// TIA Portal project "TestEssProtoFreia" (V13) (continued)
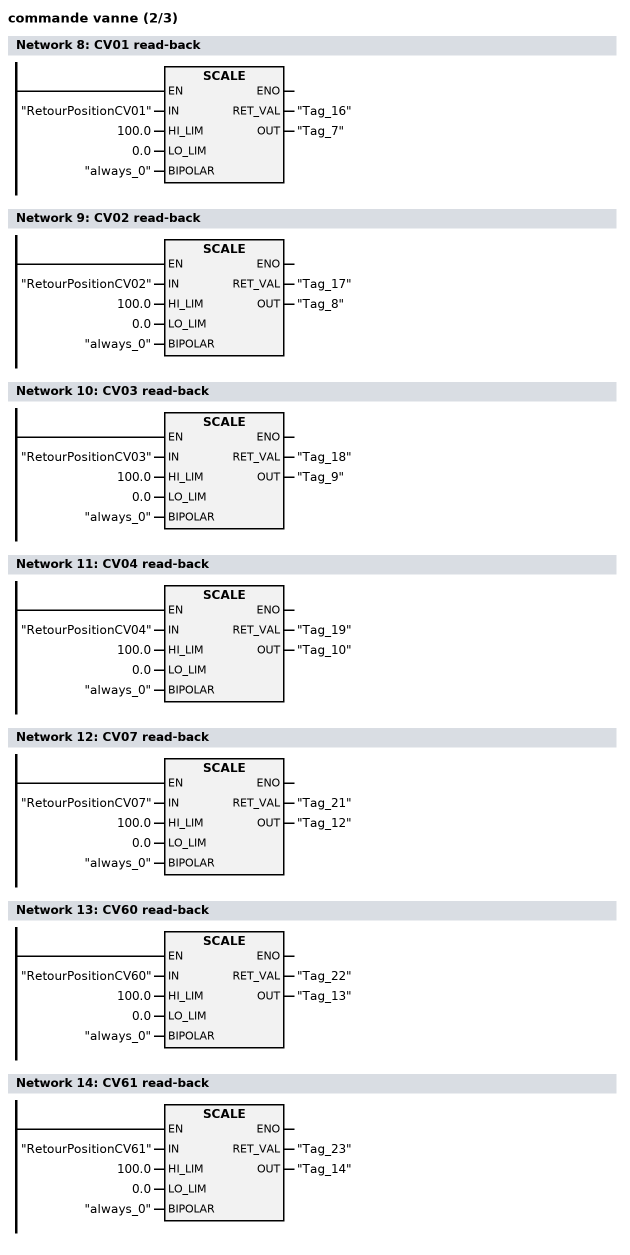
   "Tag_16" := SCALE(IN := "RetourPositionCV01",
                     HI_LIM := 100.0,
                     LO_LIM := 0.0,
                     BIPOLAR := "always_0",
                     OUT => "Tag_7");
END_REGION

REGION Network 9: CV02 read-back
   "Tag_17" := SCALE(IN := "RetourPositionCV02",
                     HI_LIM := 100.0,
                     LO_LIM := 0.0,
                     BIPOLAR := "always_0",
                     OUT => "Tag_8");
END_REGION

REGION Network 10: CV03 read-back
   "Tag_18" := SCALE(IN := "RetourPositionCV03",
                     HI_LIM := 100.0,
                     LO_LIM := 0.0,
                     BIPOLAR := "always_0",
                     OUT => "Tag_9");
END_REGION

REGION Network 11: CV04 read-back
   "Tag_19" := SCALE(IN := "RetourPositionCV04",
                     HI_LIM := 100.0,
                     LO_LIM := 0.0,
                     BIPOLAR := "always_0",
                     OUT => "Tag_10");
END_REGION

REGION Network 12: CV07 read-back
   "Tag_21" := SCALE(IN := "RetourPositionCV07",
                     HI_LIM := 100.0,
                     LO_LIM := 0.0,
                     BIPOLAR := "always_0",
                     OUT => "Tag_12");
END_REGION

REGION Network 13: CV60 read-back
   "Tag_22" := SCALE(IN := "RetourPositionCV60",
                     HI_LIM := 100.0,
                     LO_LIM := 0.0,
                     BIPOLAR := "always_0",
                     OUT => "Tag_13");
END_REGION

REGION Network 14: CV61 read-back
   "Tag_23" := SCALE(IN := "RetourPositionCV61",
                     HI_LIM := 100.0,
                     LO_LIM := 0.0,
                     BIPOLAR := "always_0",
                     OUT => "Tag_14");
END_REGION

REGION Network 15: activation PID CV03 LT03>=80%
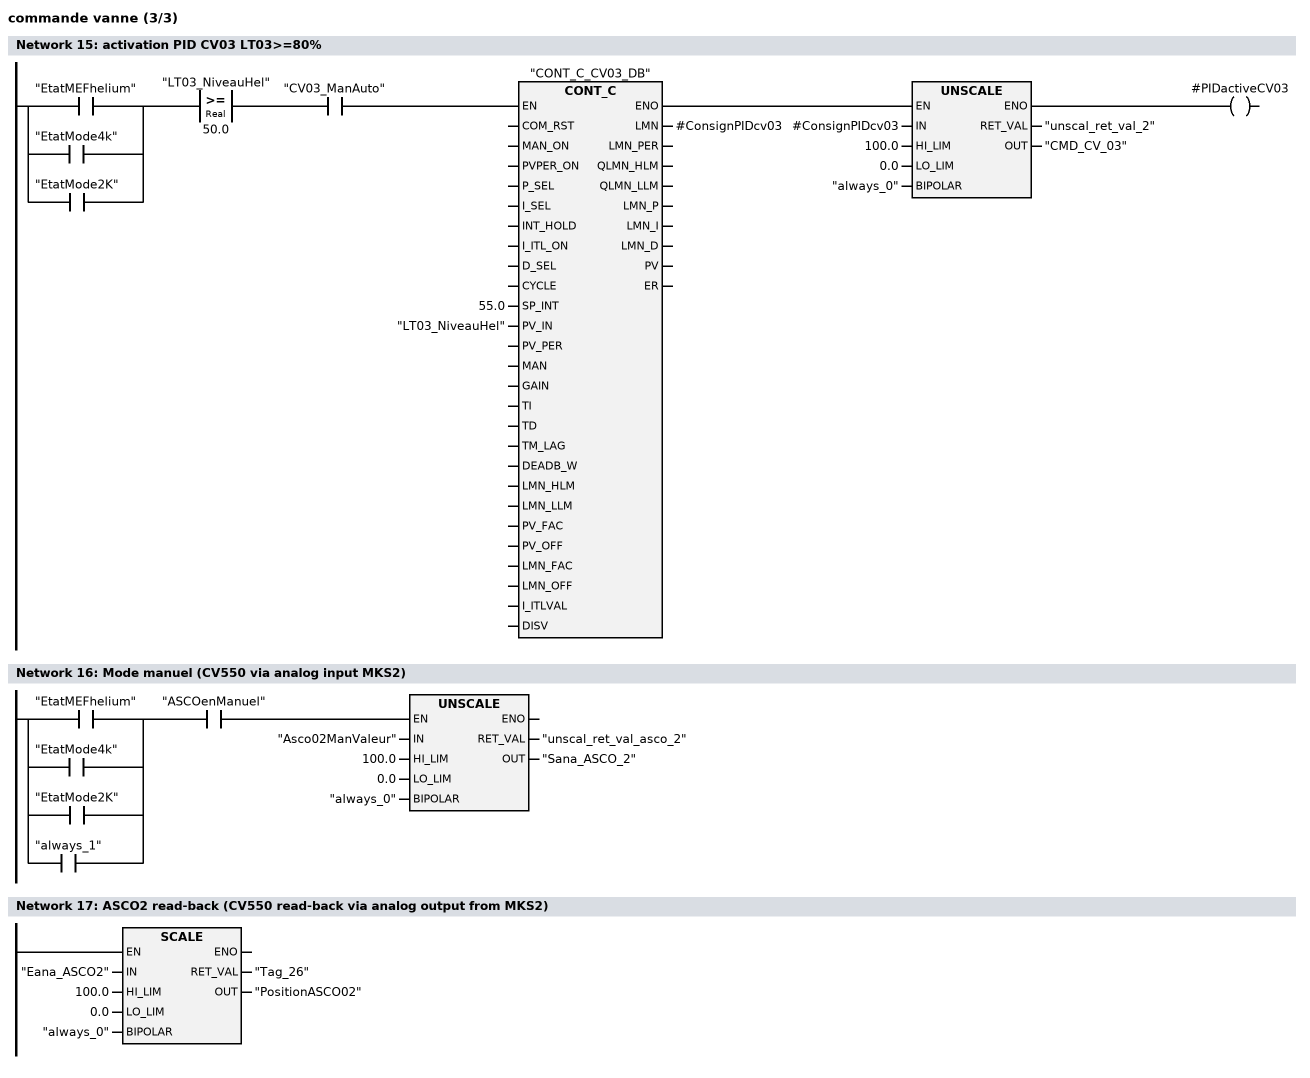
   // ENO of a box is taken as its EN; it also drops when the box reports an error
   #_w1 := ("EtatMEFhelium" OR "EtatMode4k" OR "EtatMode2K") AND ("LT03_NiveauHel" >= 50.0) AND "CV03_ManAuto";
   IF #_w1 THEN
       "CONT_C_CV03_DB"(SP_INT := 55.0, PV_IN := "LT03_NiveauHel", LMN => #ConsignPIDcv03);   // CONT_C
       "unscal_ret_val_2" := UNSCALE(IN := #ConsignPIDcv03,
                               HI_LIM := 100.0,
                               LO_LIM := 0.0,
                               BIPOLAR := "always_0",
                               OUT => "CMD_CV_03");
   END_IF;
   #PIDactiveCV03 := #_w1;
END_REGION

REGION Network 16: Mode manuel (CV550 via analog input MKS2)
   IF ("EtatMEFhelium" OR "EtatMode4k" OR "EtatMode2K" OR "always_1") AND "ASCOenManuel" THEN
       "unscal_ret_val_asco_2" := UNSCALE(IN := "Asco02ManValeur",
                               HI_LIM := 100.0,
                               LO_LIM := 0.0,
                               BIPOLAR := "always_0",
                               OUT => "Sana_ASCO_2");
   END_IF;
END_REGION

REGION Network 17: ASCO2 read-back (CV550 read-back via analog output from MKS2)
   "Tag_26" := SCALE(IN := "Eana_ASCO2",
                     HI_LIM := 100.0,
                     LO_LIM := 0.0,
                     BIPOLAR := "always_0",
                     OUT => "PositionASCO02");
END_REGION
END_FUNCTION

FUNCTION "NIveau Helium&Pression&vide" : Void   // FC2, LAD
{ S7_Optimized_Access := 'FALSE' }
VERSION : 0.1
BEGIN

REGION Network 1 (STL): scale niveau helieum LT03
         A     "always_1";
         =     #tmpb;
         BLD   103;
         CALL  "FC10=SCALE"
         ( INPUT       := "Eana_NiveauH_LT03",
           VAL_MAXI    := 74.0,
           VAL_MINI    := 0.0,
           ET_MAX      := 27648,
           ET_MIN      := 0,
           Type_Entree := 0,
           PV_SEUILH   := 100.0,
           PV_SEUILB   := 0.0,
           ACQ         := #tmpb,
           ANIM        := "LT03_TypeDef",
           PV_HIGH     := "LT03_ValMax",
           PV_LOW      := "LT03_ValMin",
           PV          := "LT03_NiveauHel",
           ALM_HIGH    := "LT03_DepHaut",
           ALM_LOW     := "LT03_DepBas",
           ALM_SENSOR  := "LT03_DefSond"
         );
         NOP   0;
END_REGION

REGION Network 2 (STL): Copy LT03 to Epics
         L     "LT03_NiveauHel";
         T     "PLC_to_Epics".LT03.Level;
         L     "LT03_TypeDef";
         T     "PLC_to_Epics".LT03.Visu;
         A     "LT03_DefSond";
         =     "PLC_to_Epics".LT03.SensorFlt;
         A     "LT03_DepHaut";
         =     "PLC_to_Epics".LT03.OverRange;
         A     "LT03_DepBas";
         =     "PLC_to_Epics".LT03.UnderRange;
END_REGION

REGION Network 3 (STL): scale niveau helieum LT01
         A     "always_1";
         =     #tmpb;
         BLD   103;
         CALL  "FC10=SCALE"
         ( INPUT       := "Eana_NiveauH_LT01",
           VAL_MAXI    := 74.0,
           VAL_MINI    := 0.0,
           ET_MAX      := 27648,
           ET_MIN      := 0,
           Type_Entree := 0,
           PV_SEUILH   := 100.0,
           PV_SEUILB   := 0.0,
           ACQ         := #tmpb,
           ANIM        := "LT01_TypeDef",
           PV_HIGH     := "LT01_ValMax",
           PV_LOW      := "LT01_ValMin",
           PV          := "LT01_NiveauHel",
           ALM_HIGH    := "LT01_DepHaut",
           ALM_LOW     := "LT01_DepBas",
           ALM_SENSOR  := "LT01_DefSond"
         );
         NOP   0;
END_REGION

REGION Network 4 (STL): Copy LT01 to Epics
         L     "LT01_NiveauHel";
         T     "PLC_to_Epics".LT01.Level;
         L     "LT01_TypeDef";
         T     "PLC_to_Epics".LT01.Visu;
         A     "LT01_DefSond";
         =     "PLC_to_Epics".LT01.SensorFlt;
         A     "LT01_DepHaut";
         =     "PLC_to_Epics".LT01.OverRange;
         A     "LT01_DepBas";
         =     "PLC_to_Epics".LT01.UnderRange;
END_REGION

REGION Network 5: Set an interlock signal for RF slow interlock
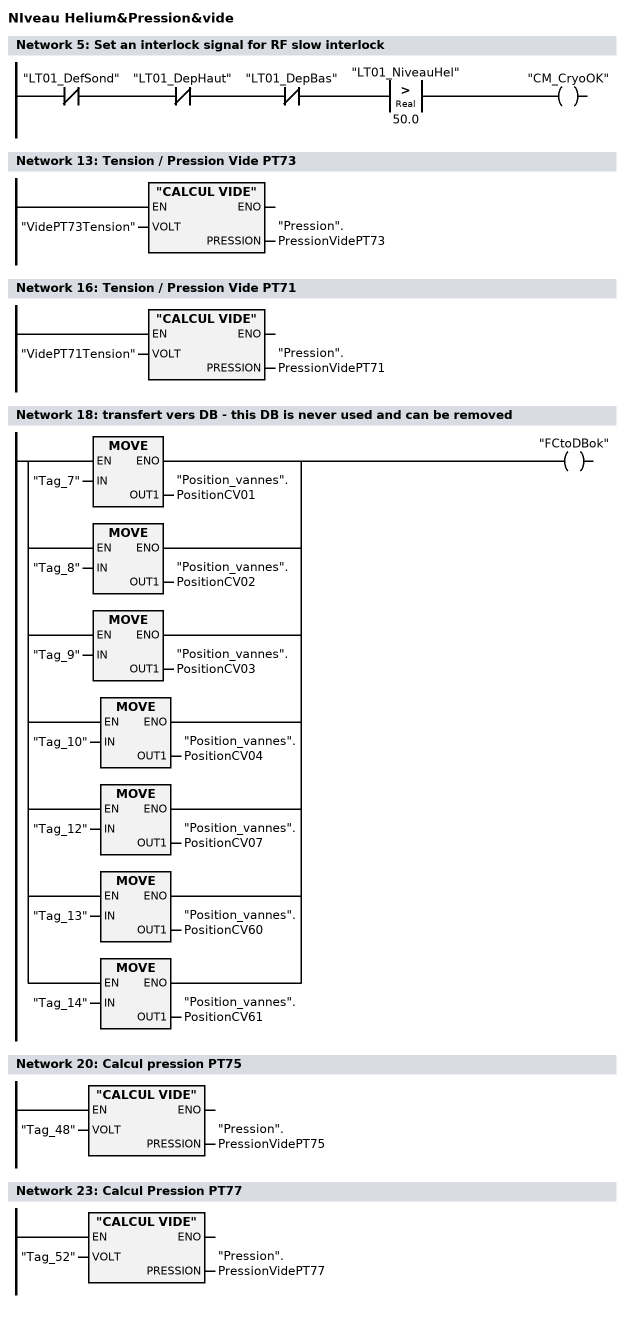
   RUNG wire#powerrail
      I_Contact( "LT01_DefSond" )
      I_Contact( "LT01_DepHaut" )
      I_Contact( "LT01_DepBas" )
      { S7_Templates := "SrcType := Real" } GT_Contact(in1 := "LT01_NiveauHel", in2 := 50.0)
      Coil( "CM_CryoOK" )
   END_RUNG
   // the same network as SCL:
   "CM_CryoOK" := NOT "LT01_DefSond" AND NOT "LT01_DepHaut" AND NOT "LT01_DepBas" AND ("LT01_NiveauHel" > 50.0);
END_REGION

REGION Network 6 (STL): scale pression PT60 ecran thermique
         A     "always_0";
         =     #tmpb;
         BLD   103;
         CALL  SCALE
         ( IN      := "Eana_PressionPT60",
           HI_LIM  := 2660.0,
           LO_LIM  := 0.0,
           BIPOLAR := #tmpb,
           RET_VAL := "ScaleErreurPT60",
           OUT     := "Pression".PressionPT60_Val
         );
         NOP   0;
END_REGION

REGION Network 7 (STL): Copy PT60 to Epics
         L     "Pression".PressionPT60_Val;
         T     "PLC_to_Epics".PT60;
END_REGION

REGION Network 8 (STL): scale pression PT01
         A     "always_0";
         =     #tmpb;
         BLD   103;
         CALL  SCALE
         ( IN      := "Eana_PressionPT01",
           HI_LIM  := 2660.0,
           LO_LIM  := 0.0,
           BIPOLAR := #tmpb,
           RET_VAL := "ScaleErreurPT01",
           OUT     := "Pression".PressionPT01_Val
         );
         NOP   0;
END_REGION

REGION Network 9 (STL): Copy PT01 to Epics
         L     "Pression".PressionPT01_Val;
         T     "PLC_to_Epics".PT01;
END_REGION

REGION Network 10 (STL): scale pression diff
         A     "always_1";
         =     #tmpb;
         BLD   103;
         CALL  SCALE
         ( IN      := "Eana_PressionDiff",
           HI_LIM  := 1.33322,
           LO_LIM  := -1.33322,
           BIPOLAR := #tmpb,
           RET_VAL := "ScaleErreurPressionDiff",
           OUT     := "Pression".PressionDiff
         );
         NOP   0;
END_REGION

REGION Network 11 (STL): Copy PT04 to Epics
         L     "Pression".PressionDiff;
         T     "PLC_to_Epics".PT04;
END_REGION

REGION Network 12 (STL): sclae vide VB PT73
         A     "always_0";
         =     #tmpb;
         BLD   103;
         CALL  SCALE
         ( IN      := "Eana_VidePT73",
           HI_LIM  := 10.0,
           LO_LIM  := 0.0,
           BIPOLAR := #tmpb,
           RET_VAL := "ScaleErreurVidePT73",
           OUT     := "VidePT73Tension"
         );
         NOP   0;
END_REGION

REGION Network 13: Tension / Pression Vide PT73
   RUNG wire#powerrail
      "CALCUL VIDE"(VOLT := "VidePT73Tension", PRESSION => "Pression".PressionVidePT73)
   END_RUNG
   // the same network as SCL:
   "CALCUL VIDE"(VOLT := "VidePT73Tension", PRESSION => "Pression".PressionVidePT73);
END_REGION

REGION Network 14 (STL): Copy PT73 to Epics
         L     "Pression".PressionVidePT73;
         T     "PLC_to_Epics".PT73;
END_REGION

REGION Network 15 (STL): scale vide CM PT71
         A     "always_0";
         =     #tmpb;
         BLD   103;
         CALL  SCALE
         ( IN      := "Eana_VidePT71",
           HI_LIM  := 10.0,
           LO_LIM  := 0.0,
           BIPOLAR := #tmpb,
           RET_VAL := "ScaleErreurVidePT71",
           OUT     := "VidePT71Tension"
         );
         NOP   0;
END_REGION

REGION Network 16: Tension / Pression Vide PT71
   RUNG wire#powerrail
      "CALCUL VIDE"(VOLT := "VidePT71Tension", PRESSION => "Pression".PressionVidePT71)
   END_RUNG
   // the same network as SCL:
   "CALCUL VIDE"(VOLT := "VidePT71Tension", PRESSION => "Pression".PressionVidePT71);
END_REGION

REGION Network 17 (STL): Copy PT71 to Epics
         L     "Pression".PressionVidePT71;
         T     "PLC_to_Epics".PT71;
END_REGION

REGION Network 18: transfert vers DB - this DB is never used and can be removed
   RUNG wire#powerrail
      { S7_GenerateENO := "TRUE" } Move(in := "Tag_7", out1 => "Position_vannes".PositionCV01)
      wire#w1
      Coil( "FCtoDBok" )
   END_RUNG
   RUNG wire#powerrail
      { S7_GenerateENO := "TRUE" } Move(in := "Tag_8", out1 => "Position_vannes".PositionCV02)
   END_RUNG wire#w1
   RUNG wire#powerrail
      { S7_GenerateENO := "TRUE" } Move(in := "Tag_9", out1 => "Position_vannes".PositionCV03)
   END_RUNG wire#w1
   RUNG wire#powerrail
      { S7_GenerateENO := "TRUE" } Move(in := "Tag_10", out1 => "Position_vannes".PositionCV04)
   END_RUNG wire#w1
   RUNG wire#powerrail
      { S7_GenerateENO := "TRUE" } Move(in := "Tag_12", out1 => "Position_vannes".PositionCV07)
   END_RUNG wire#w1
   RUNG wire#powerrail
      { S7_GenerateENO := "TRUE" } Move(in := "Tag_13", out1 => "Position_vannes".PositionCV60)
   END_RUNG wire#w1
   RUNG wire#powerrail
      { S7_GenerateENO := "TRUE" } Move(in := "Tag_14", out1 => "Position_vannes".PositionCV61)
   END_RUNG wire#w1
   // the same network as SCL:
   // ENO of a box is taken as its EN; it also drops when the box reports an error
   "Position_vannes".PositionCV01 := "Tag_7";
   "Position_vannes".PositionCV02 := "Tag_8";
   "Position_vannes".PositionCV03 := "Tag_9";
   "Position_vannes".PositionCV04 := "Tag_10";
   "Position_vannes".PositionCV07 := "Tag_12";
   "Position_vannes".PositionCV60 := "Tag_13";
   "Position_vannes".PositionCV61 := "Tag_14";
   "FCtoDBok" := TRUE OR TRUE OR TRUE OR TRUE OR TRUE OR TRUE OR TRUE;
END_REGION

REGION Network 19 (STL): Scale vide PT75
         A     "always_0";
         =     #tmpb;
         BLD   103;
         CALL  SCALE
         ( IN      := "Eana_VidePT75",
           HI_LIM  := 10.0,
           LO_LIM  := 0.0,
           BIPOLAR := #tmpb,
           RET_VAL := "Tag_50",
           OUT     := "Tag_48"
         );
         NOP   0;
END_REGION

REGION Network 20: Calcul pression PT75
   RUNG wire#powerrail
      "CALCUL VIDE"(VOLT := "Tag_48", PRESSION => "Pression".PressionVidePT75)
   END_RUNG
   // the same network as SCL:
   "CALCUL VIDE"(VOLT := "Tag_48", PRESSION => "Pression".PressionVidePT75);
END_REGION

REGION Network 21 (STL): Copy PT75 to Epics
         L     "Pression".PressionVidePT75;
         T     "PLC_to_Epics".PT75;
END_REGION

REGION Network 22 (STL): scale PT77
         A     "always_0";
         =     #tmpb;
         BLD   103;
         CALL  SCALE
         ( IN      := "Eana_VidePT77",
           HI_LIM  := 10.0,
           LO_LIM  := 0.0,
           BIPOLAR := #tmpb,
           RET_VAL := "Tag_51",
           OUT     := "Tag_52"
         );
         NOP   0;
END_REGION

REGION Network 23: Calcul Pression PT77
   RUNG wire#powerrail
      "CALCUL VIDE"(VOLT := "Tag_52", PRESSION => "Pression".PressionVidePT77)
   END_RUNG
   // the same network as SCL:
   "CALCUL VIDE"(VOLT := "Tag_52", PRESSION => "Pression".PressionVidePT77);
END_REGION

REGION Network 24 (STL): Copy PT77 to Epics
         L     "Pression".PressionVidePT77;
         T     "PLC_to_Epics".PT77;
END_REGION

REGION Network 25 (STL): FT11 - scale and copy to Epics
         A     "always_1";
         =     #tmpb;
         BLD   103;
         CALL  "FC10=SCALE"
         ( INPUT       := "FT11",
           VAL_MAXI    := 150.0,
           VAL_MINI    := -0.542534,
           ET_MAX      := 27648,
           ET_MIN      := -100,
           Type_Entree := 0,
           PV_SEUILH   := 150.0,
           PV_SEUILB   := -0.5,
           ACQ         := #tmpb,
           ANIM        := "PLC_to_Epics".FT11.Visu,
           PV_HIGH     := #tmpr,
           PV_LOW      := #tmpr,
           PV          := "PLC_to_Epics".FT11.Level,
           ALM_HIGH    := "PLC_to_Epics".FT11.OverRange,
           ALM_LOW     := "PLC_to_Epics".FT11.UnderRange,
           ALM_SENSOR  := "PLC_to_Epics".FT11.SensorFlt
         );

         NOP   0;
END_REGION

REGION Network 26 (STL): FT21 - scale and copy to Epics
         A     "always_1";
         =     #tmpb;
         BLD   103;
         CALL  "FC10=SCALE"
         ( INPUT       := "FT21",
           VAL_MAXI    := 150.0,
           VAL_MINI    := -0.542534,
           ET_MAX      := 27648,
           ET_MIN      := -100,
           Type_Entree := 0,
           PV_SEUILH   := 150.0,
           PV_SEUILB   := -0.5,
           ACQ         := #tmpb,
           ANIM        := "PLC_to_Epics".FT21.Visu,
           PV_HIGH     := #tmpr,
           PV_LOW      := #tmpr,
           PV          := "PLC_to_Epics".FT21.Level,
           ALM_HIGH    := "PLC_to_Epics".FT21.OverRange,
           ALM_LOW     := "PLC_to_Epics".FT21.UnderRange,
           ALM_SENSOR  := "PLC_to_Epics".FT21.SensorFlt
         );
         NOP   0;
END_REGION

REGION Network 27 (STL): TT102 - scale and copy to Epics
         A     "always_1";
         =     #tmpb;
         BLD   103;
         CALL  "FC10=SCALE"
         ( INPUT       := "TT102",
           VAL_MAXI    := 373.15,
           VAL_MINI    := 93.15,
           ET_MAX      := 27648,
           ET_MIN      := 0,
           Type_Entree := 0,
           PV_SEUILH   := 373.15,
           PV_SEUILB   := 93.15,
           ACQ         := #tmpb,
           ANIM        := "PLC_to_Epics".TT102.Visu,
           PV_HIGH     := #tmpr,
           PV_LOW      := #tmpr,
           PV          := "PLC_to_Epics".TT102.Level,
           ALM_HIGH    := "PLC_to_Epics".TT102.OverRange,
           ALM_LOW     := "PLC_to_Epics".TT102.UnderRange,
           ALM_SENSOR  := "PLC_to_Epics".TT102.SensorFlt
         );
         NOP   0;
END_REGION

REGION Network 28 (STL): TT202 - scale and copy to Epics
         A     "always_1";
         =     #tmpb;
         BLD   103;
         CALL  "FC10=SCALE"
         ( INPUT       := "TT202",
           VAL_MAXI    := 373.15,
           VAL_MINI    := 93.15,
           ET_MAX      := 27648,
           ET_MIN      := 0,
           Type_Entree := 0,
           PV_SEUILH   := 373.15,
           PV_SEUILB   := 93.15,
           ACQ         := #tmpb,
           ANIM        := "PLC_to_Epics".TT202.Visu,
           PV_HIGH     := #tmpr,
           PV_LOW      := #tmpr,
           PV          := "PLC_to_Epics".TT202.Level,
           ALM_HIGH    := "PLC_to_Epics".TT202.OverRange,
           ALM_LOW     := "PLC_to_Epics".TT202.UnderRange,
           ALM_SENSOR  := "PLC_to_Epics".TT202.SensorFlt
         );
         NOP   0;
END_REGION
END_FUNCTION

FUNCTION "ACQ_CABTF" : Void   // FC3, STL
{ S7_Optimized_Access := 'FALSE' }
VERSION : 0.1
BEGIN

REGION Network 1: Copie valeurs du cabtf
         CALL  BLKMOV
         ( SRCBLK  := P#I500.0 WORD 68,
           RET_VAL := #Fault_de_la_Copie,
           DSTBLK  := "VB00-LC05".CABTF
         );
         NOP   0;
END_REGION

REGION Network 2: Copy data from CATBF1 to Epics
         CALL  BLKMOV
         ( SRCBLK  := P#I518.0 WORD 16,
           RET_VAL := #Fault_de_la_Copie,
           DSTBLK  := "PLC_to_Epics".CABTF1.board1
         );
         CALL  BLKMOV
         ( SRCBLK  := P#I582.0 WORD 16,
           RET_VAL := #Fault_de_la_Copie,
           DSTBLK  := "PLC_to_Epics".CABTF1.board2
         );
         CALL  BLKMOV
         ( SRCBLK  := P#I646.0 WORD 4,
           RET_VAL := #Fault_de_la_Copie,
           DSTBLK  := "PLC_to_Epics".CABTF1.stat
         );
END_REGION

REGION Network 3: Copy data from CATBF4 to Epics
         CALL  BLKMOV
         ( SRCBLK  := P#I844.0 WORD 16,
           RET_VAL := #Fault_de_la_Copie,
           DSTBLK  := "PLC_to_Epics".CABTF4.board1
         );
         CALL  BLKMOV
         ( SRCBLK  := P#I908.0 WORD 16,
           RET_VAL := #Fault_de_la_Copie,
           DSTBLK  := "PLC_to_Epics".CABTF4.board2
         );
         CALL  BLKMOV
         ( SRCBLK  := P#I480.0 WORD 4,
           RET_VAL := #Fault_de_la_Copie,
           DSTBLK  := "PLC_to_Epics".CABTF4.stat
         );
END_REGION

REGION Network 4: Copy data from CATBF2 to Epics
         CALL  BLKMOV
         ( SRCBLK  := P#I716.0 WORD 16,
           RET_VAL := #Fault_de_la_Copie,
           DSTBLK  := "PLC_to_Epics".CABTF2.board1
         );
         CALL  BLKMOV
         ( SRCBLK  := P#I780.0 WORD 16,
           RET_VAL := #Fault_de_la_Copie,
           DSTBLK  := "PLC_to_Epics".CABTF2.board2
         );
         CALL  BLKMOV
         ( SRCBLK  := P#I472.0 WORD 4,
           RET_VAL := #Fault_de_la_Copie,
           DSTBLK  := "PLC_to_Epics".CABTF2.stat
         );
END_REGION

REGION Network 5: Copy data from CATBF3 to Epics
         CALL  BLKMOV
         ( SRCBLK  := P#I336.0 WORD 32,
           RET_VAL := #Fault_de_la_Copie,
           DSTBLK  := "PLC_to_Epics".CABTF3
         );
         CALL  BLKMOV
         ( SRCBLK  := P#I400.0 WORD 16,
           RET_VAL := #Fault_de_la_Copie,
           DSTBLK  := "PLC_to_Epics".CABTF3.board2
         );
         CALL  BLKMOV
         ( SRCBLK  := P#I464.0 WORD 4,
           RET_VAL := #Fault_de_la_Copie,
           DSTBLK  := "PLC_to_Epics".CABTF3.stat
         );
END_REGION

REGION Network 6: TT_214 (used in STBY state)
         L     "TT_214";
         T     "CM00-LC02".TT_214Res;
         NOP   0;
END_REGION

REGION Network 7: TT77
         A     "always_1";
         =     #tmpb;
         BLD   103;
         CALL  "FC10=SCALE"
         ( INPUT       := "Eana_TT77_ohm",
           VAL_MAXI    := 150.0,
           VAL_MINI    := 0.0,
           ET_MAX      := 27648,
           ET_MIN      := 0,
           Type_Entree := 0,
           PV_SEUILH   := 400.0,
           PV_SEUILB   := 0.0,
           ACQ         := #tmpb,
           ANIM        := "tt77typedef",
           PV_HIGH     := "tt77max",
           PV_LOW      := "tt77min",
           PV          := "ReceivePT100"."TT77_(R)",
           ALM_HIGH    := "tt77h",
           ALM_LOW     := "tt77l",
           ALM_SENSOR  := "tt77alm"
         );
         NOP   0;
END_REGION

REGION Network 8: TT77 - convert R -> T
         CALL  "CONVERSION R/T"
         ( "RESISTANCE _OHMS" := "ReceivePT100"."TT77_(R)",
           TEMPERATURE_KELVIN := "ReceivePT100"."TT77_(K)"
         );
         NOP   0;
END_REGION

REGION Network 9: Copy TT77 to Epics
         L     "ReceivePT100"."TT77_(K)";
         T     "PLC_to_Epics".TT77.Level;
         L     "tt77typedef";
         T     "PLC_to_Epics".TT77.Visu;
         A     "tt77alm";
         =     "PLC_to_Epics".TT77.SensorFlt;
         A     "tt77h";
         =     "PLC_to_Epics".TT77.OverRange;
         A     "tt77l";
         =     "PLC_to_Epics".TT77.UnderRange;
END_REGION

REGION Network 10: TT103 - scale and fill epics buffer
         A     "always_1";
         =     #tmpb;
         BLD   103;
         CALL  "FC10=SCALE"
         ( INPUT       := "TT103",
           VAL_MAXI    := 150.0,
           VAL_MINI    := 0.0,
           ET_MAX      := 27648,
           ET_MIN      := 0,
           Type_Entree := 0,
           PV_SEUILH   := 400.0,
           PV_SEUILB   := 0.0,
           ACQ         := #tmpb,
           ANIM        := "PLC_to_Epics".TT103.Visu,
           PV_HIGH     := #tmpr,
           PV_LOW      := #tmpr,
           PV          := #resistance,
           ALM_HIGH    := "PLC_to_Epics".TT103.OverRange,
           ALM_LOW     := "PLC_to_Epics".TT103.UnderRange,
           ALM_SENSOR  := "PLC_to_Epics".TT103.SensorFlt
         );
         NOP   0;
END_REGION

REGION Network 11: TT103 - convert R -> T
         CALL  "CONVERSION R/T"
         ( "RESISTANCE _OHMS" := #resistance,
           TEMPERATURE_KELVIN := "PLC_to_Epics".TT103.Level
         );
         NOP   0;
END_REGION

REGION Network 12: TT203 - scale and fill epics buffer
         A     "always_1";
         =     #tmpb;
         BLD   103;
         CALL  "FC10=SCALE"
         ( INPUT       := "TT203",
           VAL_MAXI    := 150.0,
           VAL_MINI    := 0.0,
           ET_MAX      := 27648,
           ET_MIN      := 0,
           Type_Entree := 0,
           PV_SEUILH   := 400.0,
           PV_SEUILB   := 0.0,
           ACQ         := #tmpb,
           ANIM        := "PLC_to_Epics".TT203.Visu,
           PV_HIGH     := #tmpr,
           PV_LOW      := #tmpr,
           PV          := #resistance,
           ALM_HIGH    := "PLC_to_Epics".TT203.OverRange,
           ALM_LOW     := "PLC_to_Epics".TT203.UnderRange,
           ALM_SENSOR  := "PLC_to_Epics".TT203.SensorFlt
         );
         NOP   0;
END_REGION

REGION Network 13: TT203 - convert R -> T
         CALL  "CONVERSION R/T"
         ( "RESISTANCE _OHMS" := #resistance,
           TEMPERATURE_KELVIN := "PLC_to_Epics".TT203.Level
         );
         NOP   0;
END_REGION
END_FUNCTION

FUNCTION "CALCUL VIDE" : Void   // FC4, SCL
{ S7_Optimized_Access := 'FALSE' }
VERSION : 0.1
BEGIN

   #PRESSION := 10 ** ((1.667*#VOLT) - 11.33);
END_FUNCTION

FUNCTION "PID ASCO" : Void   // FC5, LAD
{ S7_Optimized_Access := 'FALSE' }
VERSION : 0.1
   VAR_TEMP   // added for the SCL form of the ladder/FBD networks
      _w1 : Bool;
   END_VAR
BEGIN

REGION Network 1: PID ASCO 2
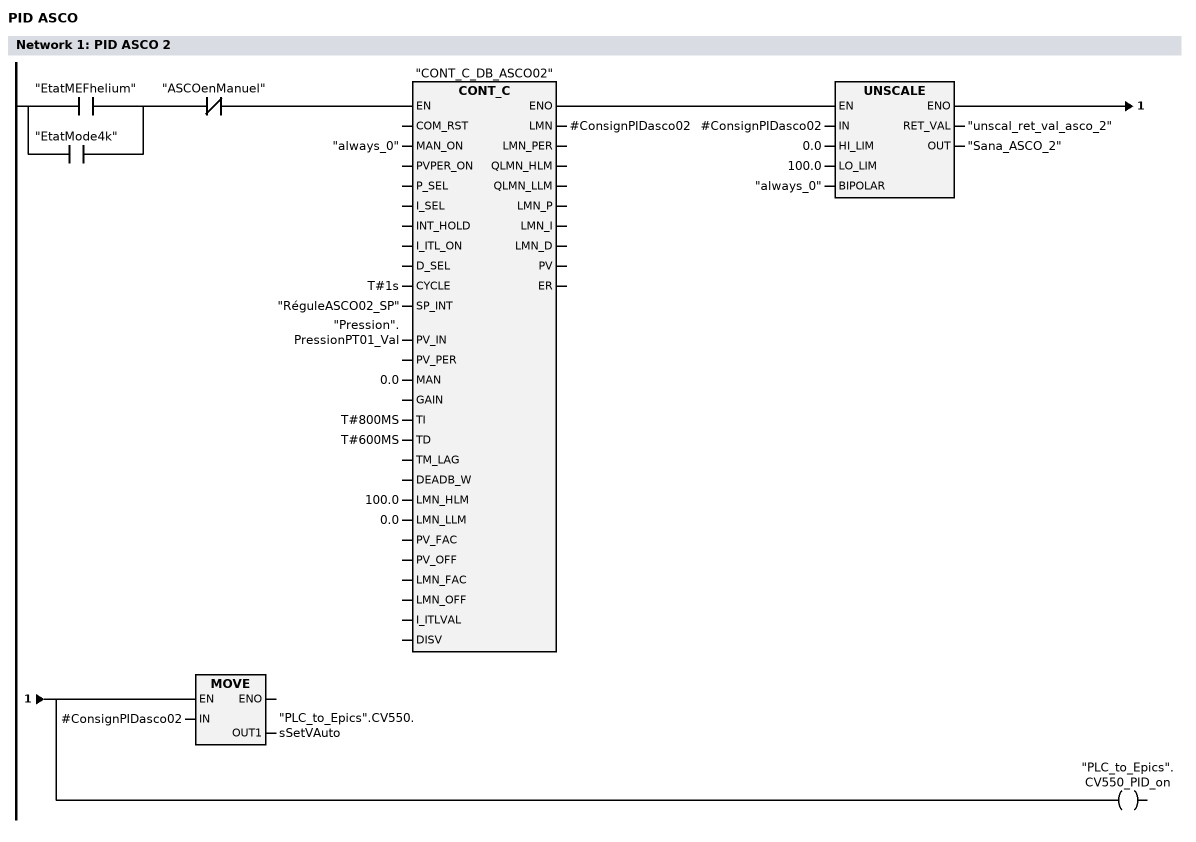
   // ENO of a box is taken as its EN; it also drops when the box reports an error
   #_w1 := ("EtatMEFhelium" OR "EtatMode4k") AND NOT "ASCOenManuel";
   IF #_w1 THEN
       "CONT_C_DB_ASCO02"(MAN_ON := "always_0",   // CONT_C
                          CYCLE := T#1s,
                          SP_INT := "RéguleASCO02_SP",
                          PV_IN := "Pression".PressionPT01_Val,
                          MAN := 0.0,
                          TI := T#800MS,
                          TD := T#600MS,
                          LMN_HLM := 100.0,
                          LMN_LLM := 0.0,
                          LMN => #ConsignPIDasco02);
       "unscal_ret_val_asco_2" := UNSCALE(IN := #ConsignPIDasco02,
                               HI_LIM := 0.0,
                               LO_LIM := 100.0,
                               BIPOLAR := "always_0",
                               OUT => "Sana_ASCO_2");
       "PLC_to_Epics".CV550.sSetVAuto := #ConsignPIDasco02;
   END_IF;
   "PLC_to_Epics".CV550_PID_on := #_w1;
END_REGION
END_FUNCTION

FUNCTION "FC10=SCALE" : Void   // FC10, FBD
TITLE = SCALE
{ S7_Optimized_Access := 'FALSE' }
VERSION : 0.1
BEGIN

REGION Network 1 (STL): input type select
         L     #Type_Entree;
         JL    LSTX;
         JU    C1;  // Valeur 0 : Tension ou courant
         JU    C2;  // Valeur 1 : PT100 en °C
         JU    C3;  // Valeur 2 : PT100 en K
   LSTX: JU    End;
END_REGION

REGION Network 2 (STL): Input type : 4-20mA, 0/10V
   // Input type  : 4-20mA, 0/10V
   // 
   // (Acquisition - Etendue mesure mini)*(Echelle max - min) + Echelle mini = mesure 
   // convertie
   // 
   // Etendue mesure maxi - mini
   C1:   L     #INPUT;
         ITD;
         DTR;
         L     #ET_MIN;
         ITD;
         DTR;
         -R;
         T     #INTER_1;  //Acquisition - etendue de mesure mini

         L     #VAL_MAXI;
         L     #VAL_MINI;
         -R;
         T     #INTER_2;  //ECHELLE MAXI - MINI

         L     #ET_MAX;
         ITD;
         DTR;
         L     #ET_MIN;
         ITD;
         DTR;
         -R;
         T     #INTER_3;  //ETENDUE DE MESURE MAXI - MINI

         L     #VAL_MINI;
         T     #INTER_4;  //ECHELLE MINI

         L     #INTER_1;
         L     #INTER_2;
         *R;
         L     #INTER_3;
         /R;
         L     #INTER_4;
         +R;
         T     #PV;
         JU    NEXT;
END_REGION

REGION Network 3 (STL): Input type : PT100 en °C
   // Input type : PT100 en °C

   C2:   L     #INPUT;
         ITD;
         DTR;
         L     10.0;
         /R;
         T     #INTER_1;



         L     #INTER_1;
         T     #PV;

         JU    NEXT;
END_REGION

REGION Network 4 (STL): Input type : PT100 en K
   // Input type  : PT100 en K

   C3:   L     #INPUT;
         ITD;
         DTR;
         L     10.0;
         /R;
         L     273.0;
         +R;
         T     #INTER_1;



         L     #INTER_1;
         T     #PV;

         JU    NEXT;
END_REGION

REGION Network 5 (STL): Depassement haut de la valeur convertie
   // Dépassement haut et bas process de la valeur
   NEXT: L     #PV;
         L     #PV_SEUILH;  //Test la valeur maximum pour le dépassement haut
         >R;
         =     #ALM_HIGH;

         L     #PV;
         L     #PV_SEUILB;  //Test la valeur minimum pour le dépassement bas
         <R;
         =     #ALM_LOW;
END_REGION

REGION Network 6 (STL): Depassement bas de la valeur convertie
   // Défaut capteur

         L     #INPUT;
         L     #ET_MAX;
         >I;
         O(;
         L     #INPUT;
         L     #ET_MIN;
         <I;
         );
         =     #ALM_TEMP;

         A     #ALM_TEMP;
         S     #ALM_SENSOR;

         AN    #ALM_TEMP;
         A     #ACQ;
         R     #ALM_SENSOR;

         NOP   0;
END_REGION

REGION Network 7 (STL): Recopie des mini et maxi de la mesure
   // Recopie des mini et maxi de la mesure
         L     #VAL_MAXI;  //Charge le maxi
         T     #PV_HIGH;

         L     #VAL_MINI;  //Charge le mini
         T     #PV_LOW;
END_REGION

REGION Network 8 (STL): Gestion du mot de défaut
   // Gestion du mot de défaut
         A     #ALM_SENSOR;
         JCN   High;  //Retourne un défaut capteur dans le mot
         L     3;  //Usually 3
         T     #ANIM;
         JU    Saut;
   High: A     #ALM_HIGH;
         JCN   Low;  //Retourne un dépassement haut dans le mot
         L     2;
         T     #ANIM;
         JU    Saut;
   Low:  A     #ALM_LOW;
         JCN   Fin;  //Retourne un dépassement bas dans le mot
         L     1;  //Usually 3
         T     #ANIM;
         JU    Saut;

   Fin:  L     0;  //Aucun défaut sur la mesure
         T     #ANIM;
   Saut: NOP   0;
END_REGION

REGION Network 9 (STL): Fin du traitement
   // Fin du traitement
   End:  NOP   0;
END_REGION
END_FUNCTION

FUNCTION "CONVERSION R/T" : Void   // FC20, SCL
{ S7_Optimized_Access := 'FALSE' }
VERSION : 0.1
BEGIN

   //#TEMPERATURE_KELVIN := REAL#29.377125832 + (REAL#2.3156100732 * #"RESISTANCE _OHMS") + (REAL#1.2102319168 * 10 ** -03 * SQR(#"RESISTANCE _OHMS"));
   #TEMPERATURE_KELVIN := REAL#29.37713 + (REAL#2.315610 * #"RESISTANCE _OHMS") + (REAL#1.210232 * 10 ** -03 * SQR(#"RESISTANCE _OHMS"));
END_FUNCTION

FUNCTION "Send_to_Epics" : Void   // FC30, LAD
{ S7_Optimized_Access := 'FALSE' }
VERSION : 0.1
   VAR_TEMP   // added for the SCL form of the ladder/FBD networks
      _w1 : Bool;
   END_VAR
BEGIN

REGION Network 1 (STL): Send timer
         AN    "EPICS_send_T1";
         L     s5t#100ms;
         SD    "EPICS_send_T0";
         A     "EPICS_send_T0";
         L     s5t#100ms;
         SD    "EPICS_send_T1";
         =     "EPICS_do_send";
END_REGION

REGION Network 2: Set ACT_SEND
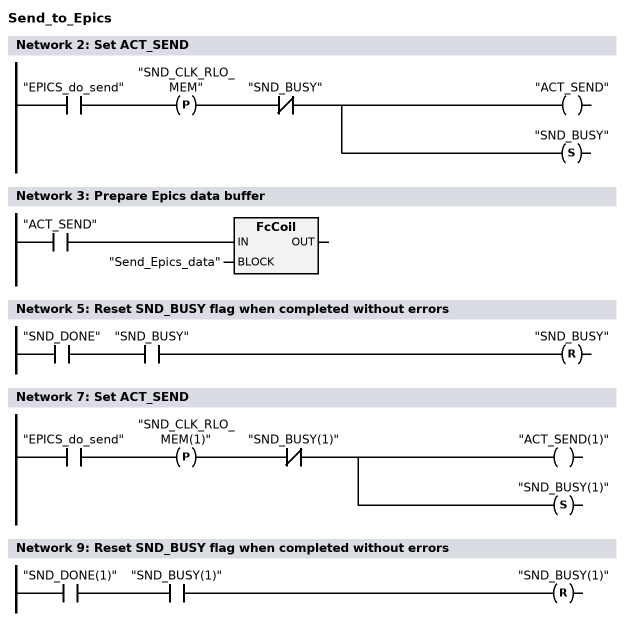
   RUNG wire#powerrail
      Contact( "EPICS_do_send" )
      P_Trig( "SND_CLK_RLO_MEM" )
      I_Contact( "SND_BUSY" )
      wire#w1
      Coil( "ACT_SEND" )
   END_RUNG
   RUNG wire#w1
      S_Coil( "SND_BUSY" )
   END_RUNG
   // the same network as SCL:
   #_w1 := "EPICS_do_send" AND NOT "SND_CLK_RLO_MEM";   // rising edge
   "SND_CLK_RLO_MEM" := "EPICS_do_send";
   "ACT_SEND" := #_w1 AND NOT "SND_BUSY";
   IF "ACT_SEND" THEN "SND_BUSY" := TRUE; END_IF;
END_REGION

REGION Network 3: Prepare Epics data buffer
   // no SCL statement known for FcCoil: written as a call
   FcCoil(block := "Send_Epics_data", in := "ACT_SEND");
END_REGION

REGION Network 4 (STL): Call AG_SEND
         CALL  AG_SEND
         ( ACT    := "ACT_SEND",
           ID     := 1,
           LADDR  := w#16#400,
           SEND   := P#DB100.DBX0.0 BYTE 2000,
           LEN    := 2000,
           DONE   := "SND_DONE",
           ERROR  := "SND_ERR",
           STATUS := "SEND_status"
         );
END_REGION

REGION Network 5: Reset SND_BUSY flag when completed without errors
   RUNG wire#powerrail
      Contact( "SND_DONE" )
      Contact( "SND_BUSY" )
      R_Coil( "SND_BUSY" )
   END_RUNG
   // the same network as SCL:
   IF "SND_DONE" AND "SND_BUSY" THEN "SND_BUSY" := FALSE; END_IF;
END_REGION

REGION Network 6 (STL): Reset SND_BUSY flag and save the status when returned error
         AN    "SND_DONE";
         A     "SND_ERR";
         JNB   ex1;
         R     "SND_BUSY";
         L     "SEND_status";
         T     "SND_STAT_SAVE";
   ex1:  NOP   0;
END_REGION

REGION Network 7: Set ACT_SEND
   RUNG wire#powerrail
      Contact( "EPICS_do_send" )
      P_Trig( "SND_CLK_RLO_MEM(1)" )
      I_Contact( "SND_BUSY(1)" )
      wire#w1
      Coil( "ACT_SEND(1)" )
   END_RUNG
   RUNG wire#w1
      S_Coil( "SND_BUSY(1)" )
   END_RUNG
   // the same network as SCL:
   #_w1 := "EPICS_do_send" AND NOT "SND_CLK_RLO_MEM(1)";   // rising edge
   "SND_CLK_RLO_MEM(1)" := "EPICS_do_send";
   "ACT_SEND(1)" := #_w1 AND NOT "SND_BUSY(1)";
   IF "ACT_SEND(1)" THEN "SND_BUSY(1)" := TRUE; END_IF;
END_REGION

REGION Network 8 (STL): Call AG_SEND
         CALL  AG_SEND
         ( ACT    := "ACT_SEND(1)",
           ID     := 2,
           LADDR  := w#16#400,
           SEND   := P#DB104.DBX0.0 BYTE 40,
           LEN    := 40,
           DONE   := "SND_DONE(1)",
           ERROR  := "SND_ERR(1)",
           STATUS := "SEND_status(1)"
         );
END_REGION

REGION Network 9: Reset SND_BUSY flag when completed without errors
   RUNG wire#powerrail
      Contact( "SND_DONE(1)" )
      Contact( "SND_BUSY(1)" )
      R_Coil( "SND_BUSY(1)" )
   END_RUNG
   // the same network as SCL:
   IF "SND_DONE(1)" AND "SND_BUSY(1)" THEN "SND_BUSY(1)" := FALSE; END_IF;
END_REGION
